(* Logix 5000 project; controller TemplateV1R0 vendor 1 type 14 code 222 rev 33.11; software revision 33.00 *)

TASK MainTask (continuous, watchdog 500 ms) : MainProgram
TASK SafetyTask (periodic, rate 20 ms, priority 10, watchdog 20 ms, safety) : SafetyProgram
TASK UnitX_XXX (event, rate 10 ms, priority 10, watchdog 500 ms) : UnitX_EMXXX

MODULES
   Local : vendor 1 type 14 code 222 (5069 0, rev 33.11)
END_MODULES

TYPE CntDescrip :
STRUCT
   ID : DINT;
   Name : STRING_16;
   Unit : STRING_08;
   Count : DINT;
   AccCount : DINT;
END_STRUCT
END_TYPE

TYPE Descriptor :
STRUCT
   ID : DINT;   // ID value of Parameter
   Name : STRING;   // Parameter name
   Unit : STRING_08;   // Unit of measure of the parameter
   Value : REAL;   // Parameter Values
END_STRUCT
END_TYPE

TYPE EquipmentModule_ModeRequest :   // Requests the equipmentmodule to switch between layers
STRUCT
   Request_Production : BOOL;   // Requests the equipmentmodule to switch between layers
   Request_Maintenance : BOOL;   // Requests the equipmentmodule to switch between layers
   Request_Manual : BOOL;   // Requests the equipmentmodule to switch between layers
   Request_Cleaning : BOOL;   // Requests the equipmentmodule to switch between layers
   Request_MES : BOOL;   // Requests the equipmentmodule to switch between layers
   Request_SemiAutomatic : BOOL;   // Requests the equipmentmodule to switch between layers
END_STRUCT
END_TYPE

TYPE EquipmentModule_SC :   // EquipmentModule- StateControl
STRUCT
   Execute_to_Completing : BOOL;   // EquipmentModule requests to move from Execute to Completing
   Unholding_to_Execute : BOOL;   // EquipmentModule requests to move from Unholding to Execute
   Starting_to_Execute : BOOL;   // EquipmentModule requests to move from Starting to Execute
   Holding_to_Held : BOOL;   // EquipmentModule requests to move from Holding to Held
   Completing_to_Completed : BOOL;   // EquipmentModule requests to move from Completing to Completed
   Suspending_to_Suspended : BOOL;   // EquipmentModule requests to move from Suspending to Suspended
   Unsuspending_to_Execute : BOOL;   // EquipmentModule requests to move from Unsuspending to Execute
   Resetting_to_Idle : BOOL;   // EquipmentModule requests to move from Resetting to Idle
   Stopping_to_Stopped : BOOL;   // EquipmentModule requests to move from Stopping to Stopped
   Clearing_to_Stopped : BOOL;   // EquipmentModule requests to move from Clearing to Stopped
   Aborting_to_Aborted : BOOL;   // EquipmentModule requests to move from Aborting to Aborted
   ons_Reset : FBD_ONESHOT;   // Reset oneshot
END_STRUCT
END_TYPE

TYPE EquipmentModule_SEQ :
STRUCT
   Clearing : DINT;   // Step nummer
   Starting : DINT;   // Step nummer
   Stopping : DINT;   // Step nummer
   Aborting : DINT;   // Step nummer
   Holding : DINT;   // Step nummer
   Unholding : DINT;   // Step nummer
   Suspending : DINT;   // Step nummer
   Unsuspending : DINT;   // Step nummer
   Resetting : DINT;   // Step nummer
   Completing : DINT;   // Step nummer
END_STRUCT
END_TYPE

TYPE Ingredients :
STRUCT
   IngredientID : DINT;
   Parameter : Descriptor[20];
END_STRUCT
END_TYPE

TYPE Interface :
STRUCT
   Number : DINT;
   ControlCmdNumber : DINT;
   CmdValue : DINT;
   RemoteInterface : Descriptor[20];
END_STRUCT
END_TYPE

TYPE PhaseStatus :   // Indicator about phase
STRUCT
   IP : BOOL;   // Phase is executing
   PC : BOOL;   // Phase complete
   EN : BOOL;   // Phase is enabled
   ER : BOOL;   // Phase faulted
   Flags : SINT;   // Phase flags
   Owner : STRING;   // Name of program who owns phase
   CurrentAction : STRING;   // Status of phase for HMI
END_STRUCT
END_TYPE

TYPE PLMs :   // Status tags are used to describe the operation of the unit machine. Status tags include state commands which describe the state transitions in the Base State Model. The status tags also include parameters and process variables which describe how the machine operates.
STRUCT
   UnitModeCurrent : DINT;   // Unit Mode in Current Use
   UnitModeRequested : BOOL;   // Requested Unit Mode Change
   UnitModeChangeInProcess : BOOL;   // Requested Unit Mode Change in Process
   StateCurrent : DINT;   // Current State Number
   StateRequested : DINT;   // Target State.
   StateChangeInProcess : BOOL;   // State Change in Process.
   MachSpeed : REAL;   // Current Machine Speed
   CurMachSpeed : REAL;   // Current Machine Speed in Primary Packages/Minute
   MaterialInterlock : BOOL;   // Materials Ready
   RemoteInterface : Interface[10];   // !!Currently not in use!! Upstream or Downstream Machine
   Parameter : Descriptor[200];   // Array of Data Type Descriptor
   Product : Product;   // The Product data type can be used for defining product and product processing parameter variables
END_STRUCT
END_TYPE

TYPE PMLc :   // Command tags are used to control the operation of the unit machine. Command tags include unit state commands which control the state transitions in the Base State Model.
STRUCT
   UnitMode : DINT;   // This value is predefined by the user/OEM, and are the desired unit modes of the machine.
   UnitModeChangeRequest : BOOL;   // When a unit mode request takes place a numerical value must be present in the Command.UnitMode tag to change the unit mode.
   MachSpeed : REAL;
   MaterialsInterlocks : BOOL;
   CntrlCmd : DINT;   // 0 Undefined 1 Reset 2 Start 3 Stop 4 Hold 5 Unhold 6 Suspend 7 Unsuspend 8 Abort 9 Clear
   CmdChangeRequest : BOOL;   // This CmdChangeRequest bit will command the machine to proceed to change the state to the target state. The tag can be used to condition when a change of state can occur. The target state will be one of the states in the base state model.
   RemoteInterface : Interface[10];   // !!Currently not in use!! Upstream or Downstream Machine
   Parameter : Descriptor[200];   // Array of Data Type Descriptor
   Product : Product[5];   // The Product data type can be used for defining product and product processing parameter variables
END_STRUCT
END_TYPE

TYPE Product :
STRUCT
   ProductID : DINT;   // Product ID
   ProcessVariables : Descriptor[30];   // Process variables include set points, limits, quality parameters, etc
   Ingredients : Ingredients[1];   // hold the information needed for the raw materials that are used by the unit machine in the processing of a particular product
END_STRUCT
END_TYPE

TYPE Settings_MinMax :
STRUCT
   Max_input : REAL;   // max value user may input
   Min_input : REAL;   // min value user may input
END_STRUCT
END_TYPE

TYPE StateCurrentTime_array :   // sub array
STRUCT
   Mode : DINT[18];
END_STRUCT
END_TYPE

TYPE STRING16 :
STRUCT
   LEN : DINT;
   DATA : SINT[16];
END_STRUCT
END_TYPE

TYPE STRING_08 :   // only 8 chars
STRUCT
   LEN : DINT;
   DATA : SINT[8];
END_STRUCT
END_TYPE

ADD_ON_INSTRUCTION AlarmGenerator   (* revision 1.0 *)
VAR_IN_OUT
   EquipmentModule : EquipmentModule; {required}
END_VAR
VAR_INPUT
   Alarm_ID : DINT; {visible}
END_VAR
VAR_IN_OUT
   Alarm_Message : STRING; {required}
END_VAR
VAR_INPUT
   Alarm_Value : REAL; {visible}
   AlarmActive : BOOL; {visible}   // Alarm is triggerd, resets automaticly once signal is turned off
END_VAR
VAR
   wrk_TimeStamp : LINT; {access None}
   alarm : BOOL; {access None}
END_VAR

ROUTINE Logic   (* structured text *)
   ////////////////////////////////////////////////////////////
   //   Copyright (c)
   //------------------------------------------------------------
   //   Routine: AlarmGenerator - Logic
   //   Author: WPI\tom.reit
   //   Created: 15-11-2022
   //------------------------------------------------------------
   //   Description:
   //
   //
   //   History:
   //
   ////////////////////////////////////////////////////////////
   GSV(WallClockTime,,CurrentValue,wrk_TimeStamp);
   
   EquipmentModule.Alarm_Local[Alarm_ID].ID				:=Alarm_ID;
   EquipmentModule.Alarm_Local[Alarm_ID].Message			:=Alarm_Message;
   EquipmentModule.Alarm_Local[Alarm_ID].TimeEvent.Date	:=wrk_TimeStamp;
   EquipmentModule.Alarm_Local[Alarm_ID].Value				:=Alarm_Value;
   
   if AlarmActive then
   	EquipmentModule.Alarm_Local_Trigger[Alarm_ID]:=1;
   else
   	EquipmentModule.Alarm_Local_Trigger[Alarm_ID]:=0;
   end_if;
   
END_ROUTINE
END_ADD_ON_INSTRUCTION

ADD_ON_INSTRUCTION AnalogOutput   (* revision 1.0 *)
VAR_INPUT
   cnf_Voltage_or_Current : BOOL; {visible}   // 0 = Voltage (0-10V) 1 = Current (4-20mA)
   cnf_HighEngineeringUnit : REAL; {visible}   // Mostlikely the card HighEngineering value
   cnf_LowEngineeringUnit : REAL; {visible}   // Mostlikely the card LowEngineering value
   cnf_Max_Output : REAL; {visible}   // Highest Voltage or Current
   cnf_Min_Output : REAL; {visible}   // Lowest Voltage or Current
   Setpoint : REAL; {required}   // requested value on outputcard
END_VAR
VAR_OUTPUT
   OutputValue : REAL; {required}   // OutputValue from scale based on userinputs sets correct value
END_VAR
VAR
   Scale_Output : SCALE; {access None}
END_VAR

ROUTINE Logic   (* structured text *)
   ////////////////////////////////////////////////////////////
   //   Copyright (c)
   //------------------------------------------------------------
   //   Routine: AnalogOutput - Logic
   //   Author: WPI\tom.reit
   //   Created: 13-1-2023
   //------------------------------------------------------------
   //   Description:
   //
   //
   //   History:
   //
   ////////////////////////////////////////////////////////////
   #region Setup
   	/* Prevent user from not entering any values, if no value is enterd use the default values from the cards respectfully. */
   	if (cnf_HighEngineeringUnit = 0 AND cnf_LowEngineeringUnit = 0) then
   				/* Voltage 0-10V */
   		if NOT cnf_Voltage_or_Current then
   			cnf_HighEngineeringUnit		:=	10000;		// 	10mV
   			cnf_LowEngineeringUnit		:=	0;			//	0mV
   			cnf_Max_Output				:=	10.00;		//	10V
   			cnf_Min_Output				:=	00.00;		//	00V
   		end_if;
   				/* Current 4-20mA */
   		if cnf_Voltage_or_Current then
   			cnf_HighEngineeringUnit		:=	8191;		//	20mA
   			cnf_LowEngineeringUnit		:=	1638;		//	04mA
   			cnf_Max_Output				:=	20.00;		//	20mA
   			cnf_Min_Output				:=	04.00;		//	04mA
   		end_if;
   	end_if;
   #endregion
   
   SCL(Scale_Output);
   Scale_Output.In			:=	Setpoint;					//	Inputvalue(requested)
   Scale_Output.InRawMax	:=	cnf_Max_Output;	//	cnf_HighEngineeringUnit
   Scale_Output.InRawMin	:=	cnf_Min_Output;		//	cnf_LowEngineeringUnit
   Scale_Output.InEUMax	:=	cnf_HighEngineeringUnit;				//	Based on cnf_Voltage_or_Current
   Scale_Output.InEUMin	:=	cnf_LowEngineeringUnit;				//	Based on cnf_Voltage_or_Current
   OutputValue				:=	Scale_Output.Out;			//	Output value eigher Voltage or Current
   
END_ROUTINE
END_ADD_ON_INSTRUCTION

ADD_ON_INSTRUCTION CMP_PML   (* revision 1.0 *)
// StateCompare PackML
VAR_IN_OUT
   PackML : PACKMLv30; {required}
END_VAR
VAR_INPUT
   cnf_Aborting : BOOL; {visible}
   cnf_Aborted : BOOL; {visible}
   cnf_Clearing : BOOL; {visible}
   cnf_Stopping : BOOL; {visible}
   cnf_Stopped : BOOL; {visible}
   cnf_Resetting : BOOL; {visible}
   cnf_Idle : BOOL; {visible}
   cnf_Starting : BOOL; {visible}
   cnf_Execute : BOOL; {visible}
   cnf_Holding : BOOL; {visible}
   cnf_Held : BOOL; {visible}
   cnf_Unholding : BOOL; {visible}
   cnf_Suspending : BOOL; {visible}
   cnf_Suspended : BOOL; {visible}
   cnf_Unsuspending : BOOL; {visible}
   cnf_Completing : BOOL; {visible}
   cnf_Complete : BOOL; {visible}
END_VAR
VAR_OUTPUT
   Sts_Result : BOOL; {access Read Only, visible}   // indicator if machine is in correct state to passthrough
END_VAR

ROUTINE Logic   (* ladder *)
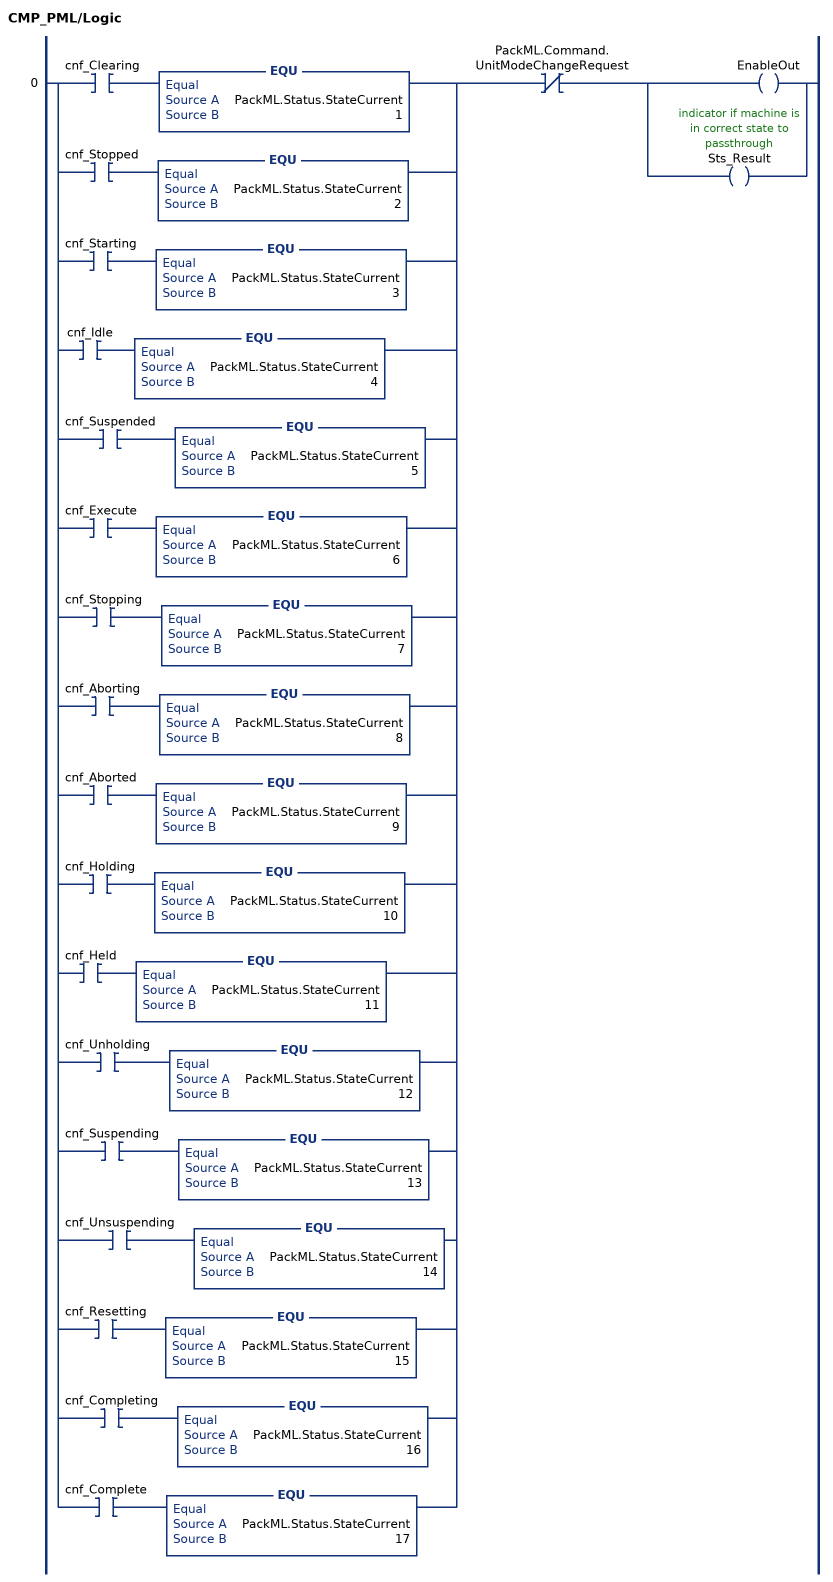
   0: [XIC(cnf_Clearing) EQU(PackML.Status.StateCurrent,1) ,XIC(cnf_Stopped) EQU(PackML.Status.StateCurrent,2) ,XIC(cnf_Starting) EQU(PackML.Status.StateCurrent,3) ,XIC(cnf_Idle) EQU(PackML.Status.StateCurrent,4) ,XIC(cnf_Suspended) EQU(PackML.Status.StateCurrent,5) ,XIC(cnf_Execute) EQU(PackML.Status.StateCurrent,6) ,XIC(cnf_Stopping) EQU(PackML.Status.StateCurrent,7) ,XIC(cnf_Aborting) EQU(PackML.Status.StateCurrent,8) ,XIC(cnf_Aborted) EQU(PackML.Status.StateCurrent,9) ,XIC(cnf_Holding) EQU(PackML.Status.StateCurrent,10) ,XIC(cnf_Held) EQU(PackML.Status.StateCurrent,11) ,XIC(cnf_Unholding) EQU(PackML.Status.StateCurrent,12) ,XIC(cnf_Suspending) EQU(PackML.Status.StateCurrent,13) ,XIC(cnf_Unsuspending) EQU(PackML.Status.StateCurrent,14) ,XIC(cnf_Resetting) EQU(PackML.Status.StateCurrent,15) ,XIC(cnf_Completing) EQU(PackML.Status.StateCurrent,16) ,XIC(cnf_Complete) EQU(PackML.Status.StateCurrent,17) ]XIO(PackML.Command.UnitModeChangeRequest)[OTE(EnableOut) ,OTE(Sts_Result) ];
END_ROUTINE
END_ADD_ON_INSTRUCTION

ADD_ON_INSTRUCTION CREATE_MERKER   (* revision 1.0 *)
VAR_INPUT
   INPUT : BOOL := 1; {required}
   RESET : BOOL; {required}
END_VAR
VAR_OUTPUT
   MERKER : BOOL; {access Read Only, visible}
END_VAR
VAR_INPUT
   I_NORMALY_OPEN : BOOL; {required}
END_VAR

ROUTINE Logic   (* ladder *)
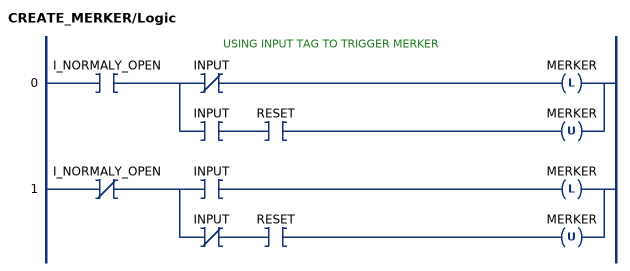
   // USING INPUT TAG TO TRIGGER MERKER
   0: XIC(I_NORMALY_OPEN)[XIO(INPUT) OTL(MERKER) ,XIC(INPUT) XIC(RESET) OTU(MERKER) ];
   1: XIO(I_NORMALY_OPEN)[XIC(INPUT) OTL(MERKER) ,XIO(INPUT) XIC(RESET) OTU(MERKER) ];
END_ROUTINE
END_ADD_ON_INSTRUCTION

ADD_ON_INSTRUCTION FLIP_FLOP   (* revision 1.0 *)
VAR_INPUT
   input_time : DINT := 1500;
END_VAR
VAR_OUTPUT
   Q : BOOL; {access Read Only, visible}
   QB : BOOL; {access Read Only, visible}
END_VAR
VAR_INPUT
   INPUT_TIME_Q : DINT; {required}   // the time Q is going to be active
   INPUT_TIME_QB : DINT; {required}   // the time QB is going to be active
END_VAR
VAR
   FLIPFLOP_TIME : DINT; {access None}
   FLIPFLOP_timer1 : TIMER; {access None}
   FLIPFLOP_timer2 : TIMER := (PRE := 7500); {access None}
   FLIPFLOP_TIME1 : DINT; {access None}
   FLIPFLOP_TIME2 : DINT; {access None}
END_VAR

ROUTINE Logic   (* ladder *)
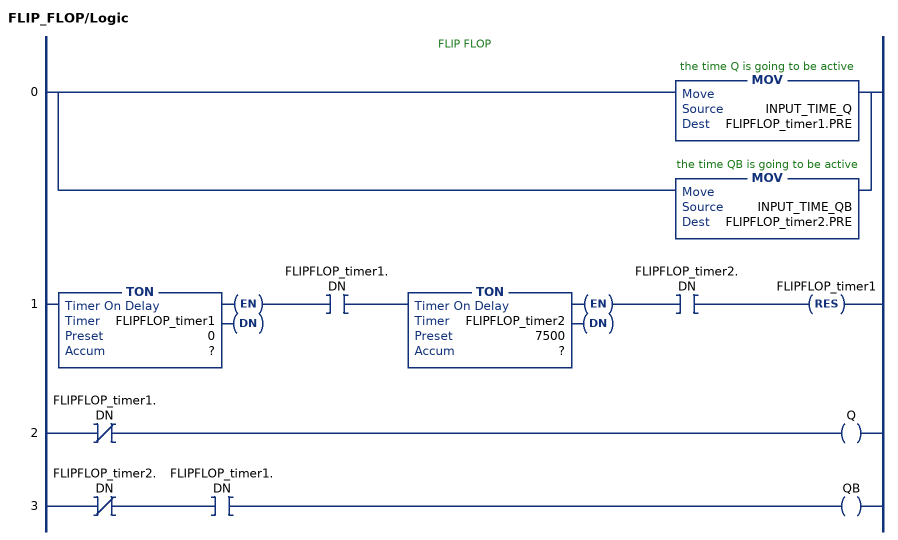
   // FLIP FLOP
   0: [MOV(INPUT_TIME_Q,FLIPFLOP_timer1.PRE) ,MOV(INPUT_TIME_QB,FLIPFLOP_timer2.PRE) ];
   1: TON(FLIPFLOP_timer1,?,?)XIC(FLIPFLOP_timer1.DN)TON(FLIPFLOP_timer2,?,?)XIC(FLIPFLOP_timer2.DN)RES(FLIPFLOP_timer1);
   2: XIO(FLIPFLOP_timer1.DN)OTE(Q);
   3: XIO(FLIPFLOP_timer2.DN)XIC(FLIPFLOP_timer1.DN)OTE(QB);
END_ROUTINE
END_ADD_ON_INSTRUCTION

ADD_ON_INSTRUCTION FLIP_FLOP_ADVANCED   (* revision 1.0 *)
VAR_OUTPUT
   Q : BOOL; {access Read Only, visible}   // Output
   QB : BOOL; {access Read Only, visible}   // Output
END_VAR
VAR_INPUT
   INPUT_HOLDING_TIME_Q : DINT; {required}   // this is the time Q will be hold after clock pulse
   INPUT_HOLDING_TIME_QB : DINT; {required}   // this is the time Q will be hold after clock pulse
   INPUT_TIME_Q : DINT := 5000; {required}
   INPUT_TIME_QB : DINT := 5000; {required}
   reset : BOOL; {required}   // this resets the Q & QB
END_VAR
VAR
   FLIPFLOP_timer1 : TIMER := (PRE := 7500); {access None}
   FLIPFLOP_timer2 : TIMER := (PRE := 7500); {access None}
   HOLDING_TIME : TIMER := (PRE := 1500); {access None}
   basic_flip_flop : FLIP_FLOP := (input_time := 1500); {access None}
   holding_timer_Q : TIMER; {access None}
   holding_timer_QB : TIMER; {access None}
   reset_ons : BOOL; {access None}
END_VAR

ROUTINE Logic   (* ladder *)
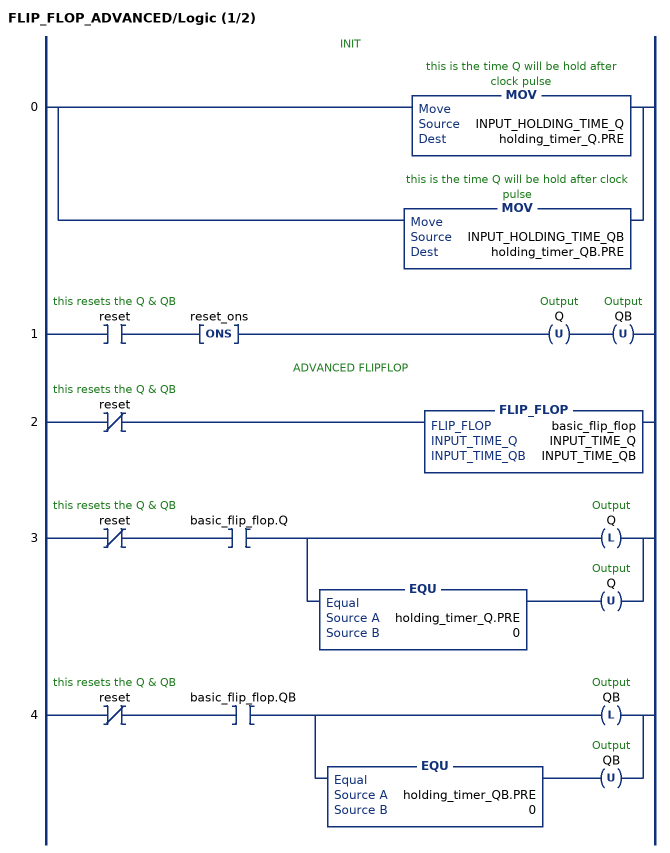
   // INIT
   0: [MOV(INPUT_HOLDING_TIME_Q,holding_timer_Q.PRE) ,MOV(INPUT_HOLDING_TIME_QB,holding_timer_QB.PRE) ];
   1: XIC(reset)ONS(reset_ons)OTU(Q)OTU(QB);
   // ADVANCED FLIPFLOP
   2: XIO(reset)FLIP_FLOP(basic_flip_flop,INPUT_TIME_Q,INPUT_TIME_QB);
   3: XIO(reset)XIC(basic_flip_flop.Q)[OTL(Q) ,EQU(holding_timer_Q.PRE,0) OTU(Q) ];
   4: XIO(reset)XIC(basic_flip_flop.QB)[OTL(QB) ,EQU(holding_timer_QB.PRE,0) OTU(QB) ];
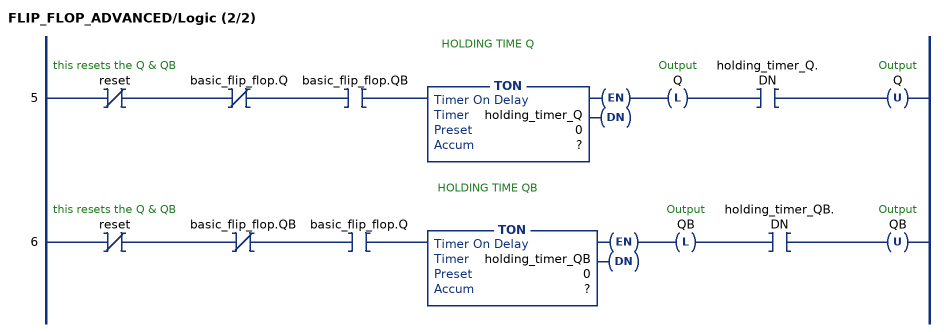
   // HOLDING TIME Q
   5: XIO(reset)XIO(basic_flip_flop.Q)XIC(basic_flip_flop.QB)TON(holding_timer_Q,?,?)OTL(Q)XIC(holding_timer_Q.DN)OTU(Q);
   // HOLDING TIME QB
   6: XIO(reset)XIO(basic_flip_flop.QB)XIC(basic_flip_flop.Q)TON(holding_timer_QB,?,?)OTL(QB)XIC(holding_timer_QB.DN)OTU(QB);
END_ROUTINE
END_ADD_ON_INSTRUCTION

ADD_ON_INSTRUCTION Generate_HMI_Tag   (* revision 1.0 *)
// Build tag for HMI
VAR_IN_OUT
   Tag : STRING; {required}
END_VAR
VAR
   Wrk_Task_Name : STRING; {access None}
   Search_String : STRING[5] := ([0] := 'unit', [1] := 'em', [2] := '_'); {access None}   // just local mem for words to find such as: Unit EM etc
   Find_pos_Unit : DINT; {access None}   // found string location
   wrk_Find_pos : DINT[5]; {access None}
   Sub_string : Substring; {access None}
   wrkTag : STRING; {access None}
   wrkTag2 : STRING; {access None}
   Wrk_Program_Name : STRING; {access None}
   Find_pos_EM : DINT; {access None}
   wrkTag3 : STRING; {access None}
   wrkTag4 : STRING; {access None}
   wrk_Insert_Pos : DINT; {access None}
END_VAR

ROUTINE Logic   (* structured text *)
// Build tag for HMI
   ////////////////////////////////////////////////////////////
   //   Copyright (c)
   //------------------------------------------------------------
   //   Routine: Generate_HMI_Tag - Logic
   //   Author: WPI\tom.reit
   //   Created: 20-12-2022
   //------------------------------------------------------------
   //   Description:
   //           Build tag for HMI
   //
   //
   //   History:
   //
   ////////////////////////////////////////////////////////////
   Search_String[0]:='unit';
   Search_String[1]:='em';
   Search_String[2]:='_';
   Search_String[3]:='t';
   Search_String[4]:='m';
   
   GSV(Task,THIS,Name,Wrk_Task_Name);					// Get task name
   LOWER(Wrk_Task_Name,Wrk_Task_Name);					// set all chars to lowercase
   FIND(Wrk_Task_Name,Search_String[0],1,Find_pos_Unit);	// search for word "unit"
   if Find_pos_Unit<>0 then
   	#region Build Unit tag
   		#region stage 1. Get UnitXXX_
   			FIND(Wrk_Task_Name,Search_String[2],Find_pos_Unit,wrk_Find_pos[1]);			// search for word "_"
   			Find_pos_Unit 		:= Find_pos_Unit 	-1;									// subtract 1 since array does not start at 1 but at 0.
   			wrk_Find_pos[1] 	:= wrk_Find_pos[1]	-0;									// subtract 0 since we need _ at the end of word.
   			Substring(Sub_string,Wrk_Task_Name,Find_pos_Unit,wrk_Find_pos[1],wrkTag);	// Set result to Tag
   		#endregion
   		#region stage 2. Get num from UnitXXX_
   			wrk_Find_pos[2]:=wrkTag.LEN;
   			FIND(wrkTag,Search_String[3],1,wrk_Find_pos[2]);						// search for word "t" used in word "unit" since after the letter t, unit nummer is expected
   			Substring(Sub_string,wrkTag,wrk_Find_pos[2],wrk_Find_pos[1],wrkTag2);	// Set result to Tag
   		#endregion
   	#endregion
   	#region Build EquipmentModule tag
   		GSV(Program,THIS,Name,Wrk_Program_Name);											// Get task name
   		LOWER(Wrk_Program_Name,Wrk_Program_Name);											// set all chars to lowercase
   		FIND(Wrk_Program_Name,Search_String[1],1,Find_pos_EM);								// search for word "em"
   		#region stage 3. Get UnitXXX_EMXXX_
   			FIND(Wrk_Program_Name,Search_String[2],Find_pos_EM,wrk_Find_pos[2]);			// search for word "_"
   			Find_pos_EM 		:= Find_pos_EM 		-1;										// subtract 1 since array does not start at 1 but at 0.
   			wrk_Find_pos[2] 	:= wrk_Find_pos[2]	-0;										// subtract 0 since we need _ at the end of word.
   			Substring(Sub_string,Wrk_Program_Name,Find_pos_EM,wrk_Find_pos[2],wrkTag3);	// Set result to Tag
   		#endregion
   		#region stage 4. Get num from EM_
   			wrk_Find_pos[3]:=wrkTag3.LEN;
   			FIND(wrkTag3,Search_String[4],1,wrk_Find_pos[4]);								// search for word "m" used in word "em" since after the letter m, unit nummer is expected
   			Substring(Sub_string,wrkTag3,wrk_Find_pos[4],wrk_Find_pos[3],wrkTag4);			// Set result to Tag
   		#endregion
   		wrk_Insert_Pos	:=wrkTag2.LEN+1;													// Move index num 1 pos
   		wrkTag4.LEN		:=wrkTag4.LEN-1;													// remove "_" from string.
   	#endregion
   	INSERT(wrkTag2,wrkTag4,wrk_Insert_Pos,Tag);											// build final string
   else
   	Tag:='XXXX';
   end_if;
   
   
   
   
END_ROUTINE
END_ADD_ON_INSTRUCTION

ADD_ON_INSTRUCTION HMI_DIG_Sensor   (* revision 1.0, vendor WPI *)
// Help:
// 0 = NO
// 1 = NC
VAR_INPUT
   NC_or_NO_Mode : BOOL; {visible}   // 0 = NC 1 = NO
   Input : BOOL; {required}
   reset : BOOL; {required}
END_VAR
VAR_OUTPUT
   Alarm : BOOL; {access Read Only, visible}
END_VAR
VAR_INPUT
   Simulatie : BOOL; {visible}
   SimulatieValue : BOOL; {visible}
END_VAR
VAR
   C_M : CREATE_MERKER := (INPUT := 1); {access None}   // Create Merker
   NC_NO : BOOL; {access None}   // Normaly open or Normaly Closed 0= NC 1 = NO
   split_char : STRING; {access None}
   Found_location : DINT; {access None}
   Num_res : DINT; {access None}
   UpperTag : STRING16; {access None}
   LowerTag : STRING16; {access None}
END_VAR

ROUTINE Logic   (* ladder *)
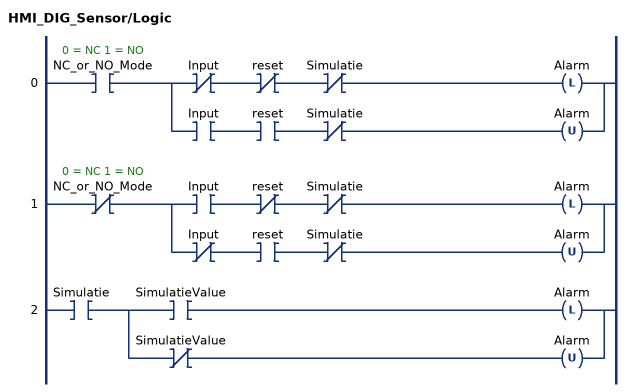
   0: XIC(NC_or_NO_Mode)[XIO(Input) XIO(reset) XIO(Simulatie) OTL(Alarm) ,XIC(Input) XIC(reset) XIO(Simulatie) OTU(Alarm) ];
   1: XIO(NC_or_NO_Mode)[XIC(Input) XIO(reset) XIO(Simulatie) OTL(Alarm) ,XIO(Input) XIC(reset) XIO(Simulatie) OTU(Alarm) ];
   2: XIC(Simulatie)[XIC(SimulatieValue) OTL(Alarm) ,XIO(SimulatieValue) OTU(Alarm) ];
END_ROUTINE
END_ADD_ON_INSTRUCTION

ADD_ON_INSTRUCTION HMI_IA_Sensor   (* revision 1.0, vendor WPI, ExecutePrescan *)
VAR_OUTPUT
   Alarm : BOOL; {visible}   // once outputvalue is not within alarmvalue low and high
END_VAR
VAR_INPUT
   AlarmValue_HIGH : REAL; {required}   // highest alarm value, based on scaled_max
   AlarmValue_LOW : REAL; {required}   // lowest alarm value based on scaled min
   InRawMax : REAL; {required}   // highest measurable value
   inRawMin : REAL; {required}   // Lowest measurable value
   Scaled_Max : REAL; {required}   // used defined Highest value (Temperature, pressure, etc)
   Scaled_Min : REAL; {required}   // used defined lowest value (Temperature, pressure, etc)
   RawSensorValue : REAL; {required}   // Sensor input from point IO card
END_VAR
VAR_OUTPUT
   OutputValue : REAL; {visible}   // scaled value
END_VAR
VAR_INPUT
   cnf_Set_100 : BOOL; {visible}   // Set inrawmax at current raw value
   cnf_Set_0 : BOOL; {visible}   // Set inrawmin at current raw value
   reset : BOOL; {required}   // Reset the alarm if alarm was true
   cnf_Use_MovingAvg : BOOL; {visible}   // 0 = no moving avg 1 = use moving avg
   MovingAvgNumberOfSamples : DINT; {visible}   // Set size of moving avg, can never be larger then array size
   MovingAvgSampleRate : DINT; {visible}   // in ms
   Simulation : BOOL; {visible}   // Set to true to bypass input rawvalue and use simulationvalue
   SimulationValue : REAL; {visible}   // Value to use for sensor once simulation is set to true
END_VAR
VAR
   HMI_Sensor : IA_SENSOR; {access None}
   Found_location : DINT; {access None}
   split_char : STRING_16; {access None}
   Num_res : DINT; {access None}
   UpperTag : STRING_16; {access None}
   LowerTag : STRING_16; {access None}
   MovingAvg : MOVING_AVERAGE := (SampleEnable := 1, NumberOfSamples := 1); {access None}
   StorageArrayMovingAvg : REAL[150]; {access None}
   wrk_arraySize : DINT; {access None}   // array size
   T_MovingAvg : FBD_TIMER; {access None}
   Build_Upper_Tag_AOI : Generate_HMI_Tag; {access None}
   Sts_Upper_Tag : STRING; {access Read Only}
   wrk_AddonName : STRING; {access None}
   GetLowerTag : Substring; {access None}
   Sts_Lower_Tag : STRING; {access Read Only}
   Sts_Show_HMIControls : BOOL;   // Show Controls
   Sts_HMI_Color : DINT; {access Read Only}   // 0 = grey 1 = green 2 = blue
END_VAR

ROUTINE Logic   (* structured text *)
   ////////////////////////////////////////////////////////////
   //   Copyright (c)
   //------------------------------------------------------------
   //   Routine: Logic
   //   Author: WPI\tom.reit
   //   Created: 31-5-2022
   //------------------------------------------------------------
   //   Description:
   //
   //
   //   History:
   //
   ////////////////////////////////////////////////////////////
   #region Read sensor value
   	#region connect input values to local addon
   		IA_SENSOR(
   					HMI_Sensor,
   					InRawMax,
   					inRawMin,
   					Scaled_Max,
   					Scaled_Min,
   					RawSensorValue,
   					1,
   					Simulation,
   					SimulationValue
   				);
   
   	#endregion
   	#region Check if value is between alarm values
   	/* for example alarmvalue_high is 10 & alarmvalue_low is 5. */
   		if HMI_Sensor.OUTPUT>AlarmValue_HIGH then
   			Alarm:=1;
   		end_if;
   		if AlarmValue_LOW>HMI_Sensor.OUTPUT then
   			Alarm:=1;
   		end_if;
   	#endregion
   	#region reset alarm
   		if Alarm AND reset then
   			Alarm:=0;
   		end_if;
   	#endregion
   #endregion
   #region Moving average
   	TONR(T_MovingAvg);
   	#region moving avg interval
   		#region set sample rate of moving avg.
   			if MovingAvgSampleRate=0 then							// no sample rate is set, this means the scantime of the PLC is the sample rate.
   				T_MovingAvg.TimerEnable:=0;							// disable timer
   				MovingAvg.In:=HMI_Sensor.OUTPUT;					// Sensor output is the moving avg input.
   				else												// Samplerate is set, so the input is based on the timer input
   				T_MovingAvg.PRE:=MovingAvgSampleRate;				// Timer pre is set by user.
   				T_MovingAvg.TimerEnable:=1;							// Enable timer
   			end_if;
   		#endregion
   		if T_MovingAvg.DN then 										// once timer is done,set copy the inputvalue to the moving avg input.
   			MovingAvg.In:=HMI_Sensor.OUTPUT;						// Sensor output is the moving avg input.
   		end_if;
   	#endregion
   	if cnf_Use_MovingAvg then
   		if HMI_Sensor.MODULE_ENABLE AND NOT Alarm then
   			MovingAvg.Initialize:=0;								// not required
   			SIZE(StorageArrayMovingAvg,0,wrk_arraySize);			// get array size, so num of samples can never be larger.
   			if MovingAvgNumberOfSamples > wrk_arraySize then MovingAvgNumberOfSamples:=wrk_arraySize; end_if;	// prevent controller faulted
   			MovingAvg.NumberOfSamples:=MovingAvgNumberOfSamples;	// set function num of samples.
   
   			/* if interval is set, then look at timer done */
   			if T_MovingAvg.TimerEnable then
   				MovingAvg.SampleEnable:=T_MovingAvg.DN;				// SampleEnable to timer enable
   			end_if;
   
   			/* if interval is not set, then bypass timer */
   			if NOT T_MovingAvg.TimerEnable then
   				MovingAvg.SampleEnable:=1;							// SampleEnable to true.
   			end_if;
   
   
   			MAVE(MovingAvg,StorageArrayMovingAvg);					// moving average function.
   			OutputValue:=MovingAvg.Out;								// Copy moving avg output to addon output.
   		else
   			OutputValue:=HMI_Sensor.OUTPUT;							// if there is an alarm in the value, move the real value to the output of the sensor addon.
   		end_if;
   	else
   		OutputValue:=HMI_Sensor.OUTPUT;								// cnf_Use_MovingAvg is not set, so use the real value form the sensor to output.(bypass moving avg)
   	end_if;
   	T_MovingAvg.Reset:=T_MovingAvg.DN;							// timer resets itself.
   #endregion
   #region Calibrate sensor
   	#region Save InRawMax
   		if cnf_Set_100 then
   			InRawMax:=HMI_Sensor.RawSensorValue;	// copy rawvalue to highest value point
   			cnf_Set_100:=0;							// set signal back to false, only run once on user input.
   		end_if;
   	#endregion
   	#region Save InRawMin
   		if cnf_Set_0 then
   			inRawMin:=HMI_Sensor.RawSensorValue;	// copy rawvalue to lowest value point
   			cnf_Set_0:=0;							// set signal back to false, only run once on user input.
   		end_if;
   	#endregion
   #endregion
   
   if s:fs then
   	Generate_HMI_Tag(Build_Upper_Tag_AOI,Sts_Upper_Tag);
   	GSV(Routine,THIS,Name,wrk_AddonName);
   	Substring(GetLowerTag,wrk_AddonName,7,wrk_AddonName.LEN,Sts_Lower_Tag);
   end_if;
   
   /* 0. Grey */
   if ( OutputValue>= Scaled_Max OR Scaled_Min >= OutputValue) AND NOT Simulation then
   	Sts_HMI_Color:=0;
   end_if;
   
   /* 1. Green */
   if (Scaled_Max >= OutputValue AND OutputValue >= Scaled_Min) AND NOT Simulation then
   	Sts_HMI_Color:=1;
   end_if;
   
   /* 2. Grey */
   if Simulation then
   	Sts_HMI_Color:=2;
   end_if;
   
END_ROUTINE

ROUTINE Prescan   (* structured text *)
// set basics
   // in scale both can never be the same, only if not valid input OR if user forgot to fillin data. lets take care of that :)
   if InRawMax=inRawMin then
   	InRawMax:=20000;
   	inRawMin:=4000;
   end_if;
   
   // in scale both can never be the same, only if not valid input OR if user forgot to fillin data. lets take care of that :)
   if Scaled_Max=Scaled_Min then
   	Scaled_Max:=100;
   	Scaled_Min:=0;
   end_if;
   
   // in scale both can never be the same, only if not valid input OR if user forgot to fillin data. lets take care of that :)
   if AlarmValue_HIGH=AlarmValue_LOW then
   	AlarmValue_HIGH:=Scaled_Max;
   	AlarmValue_LOW:=Scaled_Min;
   end_if;
   
   
END_ROUTINE
END_ADD_ON_INSTRUCTION

ADD_ON_INSTRUCTION IA_SENSOR   (* revision 2.0, vendor WPI *)
// Revision note:
// Tested by Tom Reit 25-2-2020
// Help:
// This addon instruction scales an analog input from a sensor.
// InRawMax, default: 16383 (20mA)
// InRawMin, default:  3277(4mA)
// InEUMax, max sensor value
// InEUmin, min sensor value
// RawSensorValue, this is the sensor analog input
// MODULE_ENABLE, this enables the module.
// SIMULATIE_ENABLE, if this is set to (TRUE/1) the scaling will be ignored and the OUTPUT will be the same as SIMULATIE_VALUE
VAR_INPUT
   InRawMax : REAL; {required}   // MAX analog value
   InRawMin : REAL; {required}   // MIN analog value
   InEUMax : REAL; {required}   // MAX scaled value
   InEUMin : REAL; {required}   // MIN scaled value
   RawSensorValue : REAL; {required}   // raw sensor value
   MODULE_ENABLE : BOOL; {required}   // TURNS ON THE MODULE
   SIMULATIE_ENABLE : BOOL; {required}   // Turns on the simulation and ignores the RawSensorValue
   SIMULATIE_VALUE : REAL; {required}   // Simulation value (make sure it is in the same range to achieve best preformance)
END_VAR
VAR_OUTPUT
   OUTPUT : REAL; {access Read Only, visible}   // Live Output value from the addon
END_VAR
VAR
   SCL_01 : SCALE; {access None}
   SEL_01 : SELECT; {access None}
   ScaledSensorValue : REAL;   // scaled value
   __l0578B6F82C94F046 : REAL; {access None}
   __lF2C86C86D0E4FACF : REAL; {access None}
   __lE33E53D79AF57856 : REAL; {access None}
   __l34092065E529AFDE : REAL; {access None}
   __l47628872F6E0CF0E : BOOL; {access None}
   __lB970390096686554 : REAL; {access None}
   __l80C1A40296D2D6C9 : BOOL; {access None}
   __l53AC6A8A11BDDEC1 : REAL; {access None}
   __lDC0EA55186A67465 : REAL; {access None}
   __fout9C8D1D58804E7A03 : BOOL[32]; {access None}
END_VAR

ROUTINE Logic   (* function block diagram *)
   SHEET 1
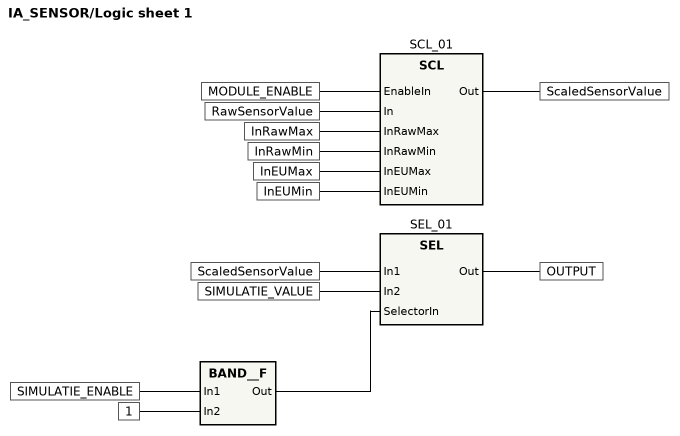
   BAND__F_1 : BAND__F(In1 := SIMULATIE_ENABLE, In2 := 1);
   SCL_01 : SCL(EnableIn := MODULE_ENABLE, In := RawSensorValue, InRawMax := InRawMax, InRawMin := InRawMin, InEUMax := InEUMax, InEUMin := InEUMin);
   SEL_01 : SEL(In1 := ScaledSensorValue, In2 := SIMULATIE_VALUE, SelectorIn := BAND__F_1.Out);
   ScaledSensorValue := SCL_01.Out;
   OUTPUT := SEL_01.Out;
END_ROUTINE
END_ADD_ON_INSTRUCTION

ADD_ON_INSTRUCTION ISA_TR_88_00_02   (* revision 1.0, ExecutePrescan *)
// Machine and Unit States:
// An Implementation Example of
// ISA-88
VAR_IN_OUT
   EMs_Status : EquipmentModule[32]; {required}   // EquipmentModules information
END_VAR
VAR_OUTPUT
   Sts_Clearing : BOOL; {access Read Only, visible}   // Clearing
   Sts_Stopped : BOOL; {access Read Only, visible}   // Stopped
   Sts_Starting : BOOL; {access Read Only, visible}   // Starting
   Sts_Idle : BOOL; {access Read Only, visible}   // Idle
   Sts_Suspended : BOOL; {access Read Only, visible}   // Suspended
   Sts_Execute : BOOL; {access Read Only, visible}   // Execute
   Sts_Stopping : BOOL; {access Read Only, visible}   // Stopping
   Sts_Aborting : BOOL; {access Read Only, visible}   // Aborting
   Sts_Aborted : BOOL; {access Read Only, visible}   // Aborted
   Sts_Holding : BOOL; {access Read Only, visible}   // Holding
   Sts_Held : BOOL; {access Read Only, visible}   // Held
   Sts_Unholding : BOOL; {access Read Only, visible}   // Unholding
   Sts_Suspending : BOOL; {access Read Only, visible}   // Suspending
   Sts_Unsuspending : BOOL; {access Read Only, visible}   // Unsuspending
   Sts_Resetting : BOOL; {access Read Only, visible}   // Resetting
   Sts_Completing : BOOL; {access Read Only, visible}   // Completing
   Sts_Complete : BOOL; {access Read Only, visible}   // Complete
   Sts_Production : BOOL; {access Read Only, visible}   // Machine is in production
   Sts_Maintenance : BOOL; {access Read Only, visible}   // Machine is in Maintenance
   Sts_Manual : BOOL; {access Read Only, visible}   // Machine is in Manual
   Sts_Cleaning : BOOL; {access Read Only, visible}   // Machine is in Cleaning
   Sts_MES : BOOL; {access Read Only, visible}   // Machine is in MES mode
   Sts_SemiAutomatic : BOOL; {access Read Only, visible}   // Machine is in Semi-Automatic
   Sts_SC_Status : UDINT; {access Read Only, visible}
END_VAR
VAR_IN_OUT
   PackTags : PACKMLv30; {required}
END_VAR
VAR_INPUT
   RecipeNumber : SINT; {visible}   // Recipe number selects which PackTag.command.product[#] will be used.
   DesignedSpeed : REAL; {visible}   // This tag represents the maximum design speed of the machine in primary packages per minute for the package configuration being run. This speed is NOT the maximum speed as specified by the manufacturer, but rather the speed the machine is designed to run in its installed environment. NOTE: In practice the maximum speed of the machine as used for efficiency calculations will be a function of how it is set up and what products it is producing.
END_VAR
VAR_OUTPUT
   Sts_MachineFaulted : BOOL; {access Read Only, visible}   // Machine recieved an fault trigger
END_VAR
VAR_INPUT
   HMI_Reset : BOOL;   // Common reset for all EMs
END_VAR
VAR
   MachineState : USINT := 255; {access None}   // Technical Report Equipment States: 1 Clearing 2 Stopped 3 Starting 4 Idle 5 Suspended 6 Execute 7 Stopping 8 Aborting 9 Aborted 10 Holding 11 Held 12 Unholding 13 Suspending 14 Unsuspending 15 Resetting 16 Completing 17 Complete
   wrk_compare_UDINT : UDINT := 65535; {access None}
   wrk_Aborting_to_Aborted : UDINT := 2#0000_0000_0000_0000_1111_1111_1111_1111; {access None}
   i : DINT; {access None}   // index num, only for local use. used for forloops
   Wrk_Aborting_to_Aborted_PC : BOOL; {access None}   // EquipmentModule(s) Aborting_to_Aborted Proces Complete
   FALSE : BOOL; {access None}   // always false
   TRUE : BOOL; {access None}   // always true
   cnf_EM_Size : DINT := 1; {access None}   // size of array for equipmentmodules
   wrk_Conversion : DINT; {access None}
   temp_sum : DINT; {access None}   // local storage
   wrk_Stopping_to_Stopped : UDINT; {access None}
   wrk_Starting_to_Execute : UDINT; {access None}
   wrk_Clearing_to_Stopped : UDINT; {access None}
   wrk_Holding_to_Held : UDINT; {access None}
   wrk_Unholding_to_Execute : UDINT; {access None}
   wrk_Suspending_to_Suspended : UDINT; {access None}
   wrk_Unsuspending_to_Execute : UDINT; {access None}
   wrk_Resetting_to_Idle : UDINT; {access None}
   wrk_Completing_to_Completed : UDINT; {access None}
   wrk_prev_state : DINT; {access None}   // local mem
   MachineMode : DINT; {access None}
   wrk_SwitchLayer_To_Cleaning : DINT; {access None}
   Feedback_Request_Cleaning : UDINT; {access None}   // local mem
   wrk_SwitchLayer_To_Maintenance : DINT; {access None}
   Feedback_Request_Maintenance : UDINT; {access None}   // local mem
   wrk_SwitchLayer_To_Manual : DINT; {access None}
   Feedback_Request_Manual : UDINT; {access None}
   wrk_SwitchLayer_To_MES : DINT; {access None}
   Feedback_Request_MES : UDINT; {access None}
   wrk_SwitchLayer_To_Production : DINT; {access None}
   Feedback_Request_Production : UDINT; {access None}
   wrk_SwitchLayer_To_SemiAutomatic : DINT; {access None}
   Feedback_Request_SemiAutomatic : UDINT; {access None}
   k : DINT; {access None}   // nested index num
   cnf_Status_RemoteInterface_ArraySize : DINT; {access None}
   ArraySize : DINT[5]; {access None}   // local array size
   wrk_RecipeNumber : DINT; {access None}   // local RecipeNum
   T_Refresh_PackTag_Status : FBD_TIMER; {access None}
   T_second_puls : FBD_TIMER; {access None}   // local timer for just 1 second
   T_Refresh_PackTag_Administration : FBD_TIMER; {access None}   // local timer
   wrk_DateTime : LINT; {access None}
   wrk_Execute_to_Completing : UDINT; {access None}
   T_ResetSignal_ON : FBD_TIMER; {access None}   // Local reset timer
   T_ResetSignal_OFF : FBD_TIMER; {access None}   // local reset timer
   T_ResetSignal_HMI : FBD_TIMER; {access None}   // reset timer from HMI
   StateHistory : StateHistory[10]; {access None}
END_VAR

ROUTINE Logic   (* structured text *)
// Machine and Unit States:
// An Implementation Example of
// ISA-88
   ////////////////////////////////////////////////////////////
   //   Copyright (c)
   //------------------------------------------------------------
   //   Routine: ISA_TR_88_00_02 - Logic
   //   Author: WPI\tom.reit
   //   Created: 2-11-2022
   //------------------------------------------------------------
   //   Description:
   //           Machine and Unit States:
   //           An Implementation Example of
   //           ISA-88
   //
   //
   //   History:
   //
   ////////////////////////////////////////////////////////////
   #region Macros / keywords
   	TRUE:=1;
   	FALSE:=0;
   	#region Second timer
   		if T_second_puls.DN then
   			T_second_puls.Reset:=TRUE;
   		else
   			T_second_puls.Reset:=FALSE;
   		end_if;
   		T_second_puls.TimerEnable	:=TRUE;
   		T_second_puls.PRE			:=1000;
   		TONR(T_second_puls);
   	#endregion
   	#region Reset timers
   	//On users request to reset or clear the machine there will be a resetSignal set for 50mS an it will be low for 100mS. once these timers are done, the machine will check feedback from EMs
   		T_ResetSignal_ON.TimerEnable	:=Sts_Clearing OR Sts_Resetting;											// once machine is in clearing or resetting or reset is pressed on HMI set reset for 50mS
   		T_ResetSignal_ON.PRE			:=50;																		// reset high time
   		T_ResetSignal_ON.Reset			:=(Sts_Stopped OR Sts_Aborted OR Sts_Idle) AND T_ResetSignal_OFF.DN;		// clear timer
   
   		T_ResetSignal_OFF.PRE			:=100;																		// time reset signal off
   		T_ResetSignal_OFF.TimerEnable	:=T_ResetSignal_ON.DN;														// start time off once time on is done.
   		T_ResetSignal_OFF.Reset			:=T_ResetSignal_OFF.DN AND NOT (Sts_Clearing OR Sts_Resetting);				// clear timer
   
   		T_ResetSignal_HMI.PRE			:=50;																		// time reset signal off
   		T_ResetSignal_HMI.TimerEnable	:=(HMI_Reset OR T_ResetSignal_HMI.TT);										// start time off once time on is done.
   		T_ResetSignal_HMI.Reset			:=T_ResetSignal_HMI.DN AND NOT HMI_Reset;															// clear timer
   
   		TONR(T_ResetSignal_ON);																						// timer object
   		TONR(T_ResetSignal_OFF);																					// timer object
   		TONR(T_ResetSignal_HMI);																					// timer object
   
   		if T_ResetSignal_ON.TT then
   			for i := 0 to cnf_EM_Size do
   				if NOT EMs_Status[i].Reset_Signal then EMs_Status[i].Reset_Signal:=TRUE; end_if;					// set reset signal for all EMs
   			end_for;
   		end_if;
   		if T_ResetSignal_OFF.TT then
   			for i := 0 to cnf_EM_Size do
   				if EMs_Status[i].Reset_Signal then EMs_Status[i].Reset_Signal:=FALSE; end_if;						// unset reset signal for all EMs
   			end_for;
   		end_if;
   
   		if T_ResetSignal_HMI.TT then
   			for i := 0 to cnf_EM_Size do
   				if NOT EMs_Status[i].Reset_Signal then EMs_Status[i].Reset_Signal:=TRUE; end_if;						// set reset signal for all EMs
   			end_for;
   		end_if;
   		if T_ResetSignal_HMI.DN then
   			for i := 0 to cnf_EM_Size do
   				if EMs_Status[i].Reset_Signal then EMs_Status[i].Reset_Signal:=FALSE; end_if;						// set reset signal for all EMs
   			end_for;
   			HMI_Reset:=FALSE;
   		end_if;
   	#endregion
   
   #endregion
   #region Prevent wrk_RecipeNumber overflow & underflow
   	wrk_RecipeNumber:=RecipeNumber;				// copy RecipeNumber to wrk_RecipeNumber to ensure program uses correct RecipeNumber and does not change midway reading.
   	wrk_RecipeNumber:=abs(wrk_RecipeNumber);	// if negative value is inserted, make sure it is positive.
   	if wrk_RecipeNumber>4 then					// if wrk_RecipeNumber is bigger then 4 set it back to 4.
   		wrk_RecipeNumber:=4;
   	end_if;
   	RecipeNumber:=wrk_RecipeNumber;				// mirror wrk_RecipeNumber to RecipeNumber if user has given wrong input
   #endregion
   #region Machine States
   /*Discription
   A State transition is defined as a passage from one state to another. Transitions between
   states will occur as a result of a local, remote, or procedural State command.
   
   
   for the SC's we use the following bit manipulation run a forloop from 0 till max array size.
   each cycle of the forloop check if EMs_Status[i]Request_SC.XXXXX is true or false.
   
   since an bool can not be directly moved into an UDINT we do some clever calculations
   (1*2)^i OR (0*2)^i this will result into an DEC value based on the BIN bit num.
   
   forexample BIN the value is 1011 this is DEC 13 if we want to convert 1011 to an DEC value we cycle through each bit using an index num. so
   
   BIT value		Index num			Calculation			Result
   	1				0				(1*2)^0					1
   	0				1				(0*2)^1					0
   	1				2				(1*2)^2					4
   	1				3				(1*2)^3					8
   
   	now we sum up result which is 1+0+4+8 = 13.
   	this way we have converted an array of bools into an UDINT. Now we can compare an UDINT with an compare value(all 32 bits to TRUE)
   */
   #region Switch layer to cleaning
   	case wrk_SwitchLayer_To_Cleaning of
   		0: // check for request
   			if PackTags.Command.UnitMode = 4 AND PackTags.Command.UnitModeChangeRequest then 									// request from HMI
   				PackTags.Status.UnitModeRequested		:=TRUE;						// request mode
   				PackTags.Status.UnitModeChangeInProcess	:=TRUE;						// changing mode
   				wrk_SwitchLayer_To_Cleaning				:=1;						// Set to next step
   			end_if;
   		1: // Set all modules in request mode
   			for i :=0  to cnf_EM_Size do											// scan through all equipmentmodules
   				EMs_Status[i].Request_Mode.Request_Cleaning:=TRUE;					// set mode change to all equipmentmodules
   			end_for;
   			wrk_SwitchLayer_To_Cleaning:=2;											// set to next step
   		2: // check for feedback
   			#region Check EquipmentModule feedback
   			temp_sum:=0;															// clear old mem
   				for i := 0 to cnf_EM_Size do										// scan from 0 till max array size
   					if EMs_Status[i].Selected then									// check if EquipmentModule is selected
   						if EMs_Status[i].Request_Mode_Feedback.Request_Cleaning then// Feedback from equipmentmodule
   							Feedback_Request_Cleaning:=(1*2**i)+temp_sum; 			// state is true. convert binary to dec value. sum= bits *2 ^ i. See https://flexiple.com/developers/decimal-to-binary-conversion
   					 	else
   							Feedback_Request_Cleaning:=(0*2**i)+temp_sum; 			// state is false. convert binary to dec value. sum= bits *2 ^ i. See https://flexiple.com/developers/decimal-to-binary-conversion
   						end_if;
   					end_if;
   					if NOT EMs_Status[i].Selected then Feedback_Request_Cleaning:=(1*2**i)+temp_sum; end_if; // module is not enabled. therfor state is always true.
   					temp_sum:=Feedback_Request_Cleaning;
   				end_for;
   				if Feedback_Request_Cleaning = wrk_compare_UDINT then				// compare to compare UDINT
   					wrk_SwitchLayer_To_Cleaning:=3;									//	next step
   				end_if;
   			#endregion
   		3: // Set unit to new mode.
   			for i := 0 to cnf_EM_Size do
   				EMs_Status[i].Request_Mode.Request_Cleaning:=FALSE;				// mode select was succesfull, remove request.
   			end_for;
   			PackTags.Status.UnitModeChangeInProcess	:=FALSE;							// changing mode done
   			PackTags.Status.UnitModeRequested		:=FALSE;							// request mode
   			PackTags.Command.UnitMode				:=0;								// unlatch signal on HMI as feedback.
   			MachineMode								:=4;								// Set machine in other layer.
   			wrk_SwitchLayer_To_Cleaning				:=0;								// reset statemodel
   		else // undefined state
   			wrk_SwitchLayer_To_Cleaning:=0;
   	end_case;
   	if wrk_SwitchLayer_To_Cleaning <> 0 AND NOT (PackTags.Command.UnitMode=4) then
   		wrk_SwitchLayer_To_Cleaning:=0; 											// reset request once signal is set back to 0 and machine did not switch layer.
   	end_if;
   #endregion